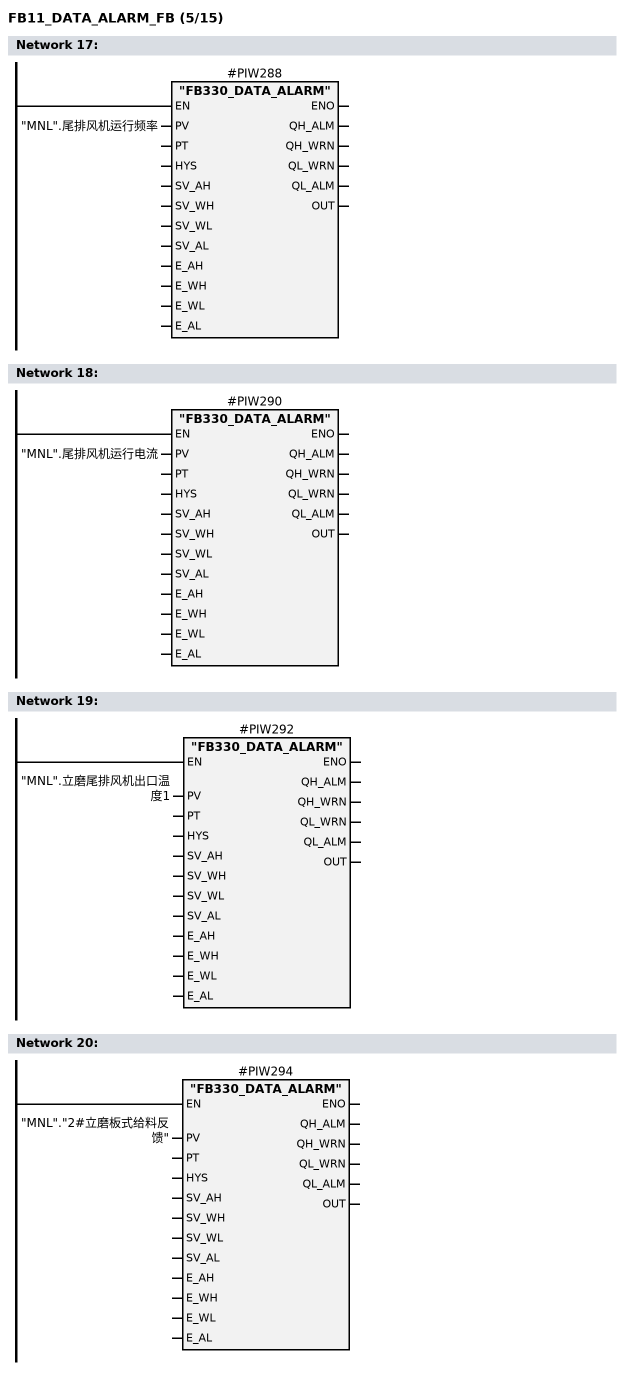
   RUNG wire#powerrail
      #PIW288(PV := "MNL".尾排风机运行频率, PT :=, HYS :=, SV_AH :=, SV_WH :=, SV_WL :=, SV_AL :=, E_AH :=, E_WH :=, E_WL :=, E_AL :=, QH_ALM =>, QH_WRN =>, QL_WRN =>, QL_ALM =>, OUT =>)
   END_RUNG
   // the same network as SCL:
   #PIW288(PV := "MNL".尾排风机运行频率);   // "FB330_DATA_ALARM"
END_REGION

REGION Network 18
   RUNG wire#powerrail
      #PIW290(PV := "MNL".尾排风机运行电流, PT :=, HYS :=, SV_AH :=, SV_WH :=, SV_WL :=, SV_AL :=, E_AH :=, E_WH :=, E_WL :=, E_AL :=, QH_ALM =>, QH_WRN =>, QL_WRN =>, QL_ALM =>, OUT =>)
   END_RUNG
   // the same network as SCL:
   #PIW290(PV := "MNL".尾排风机运行电流);   // "FB330_DATA_ALARM"
END_REGION

REGION Network 19
   RUNG wire#powerrail
      #PIW292(PV := "MNL".立磨尾排风机出口温度1, PT :=, HYS :=, SV_AH :=, SV_WH :=, SV_WL :=, SV_AL :=, E_AH :=, E_WH :=, E_WL :=, E_AL :=, QH_ALM =>, QH_WRN =>, QL_WRN =>, QL_ALM =>, OUT =>)
   END_RUNG
   // the same network as SCL:
   #PIW292(PV := "MNL".立磨尾排风机出口温度1);   // "FB330_DATA_ALARM"
END_REGION

REGION Network 20
   RUNG wire#powerrail
      #PIW294(PV := "MNL"."2#立磨板式给料反馈", PT :=, HYS :=, SV_AH :=, SV_WH :=, SV_WL :=, SV_AL :=, E_AH :=, E_WH :=, E_WL :=, E_AL :=, QH_ALM =>, QH_WRN =>, QL_WRN =>, QL_ALM =>, OUT =>)
   END_RUNG
   // the same network as SCL:
   #PIW294(PV := "MNL"."2#立磨板式给料反馈");   // "FB330_DATA_ALARM"
END_REGION

REGION Network 21
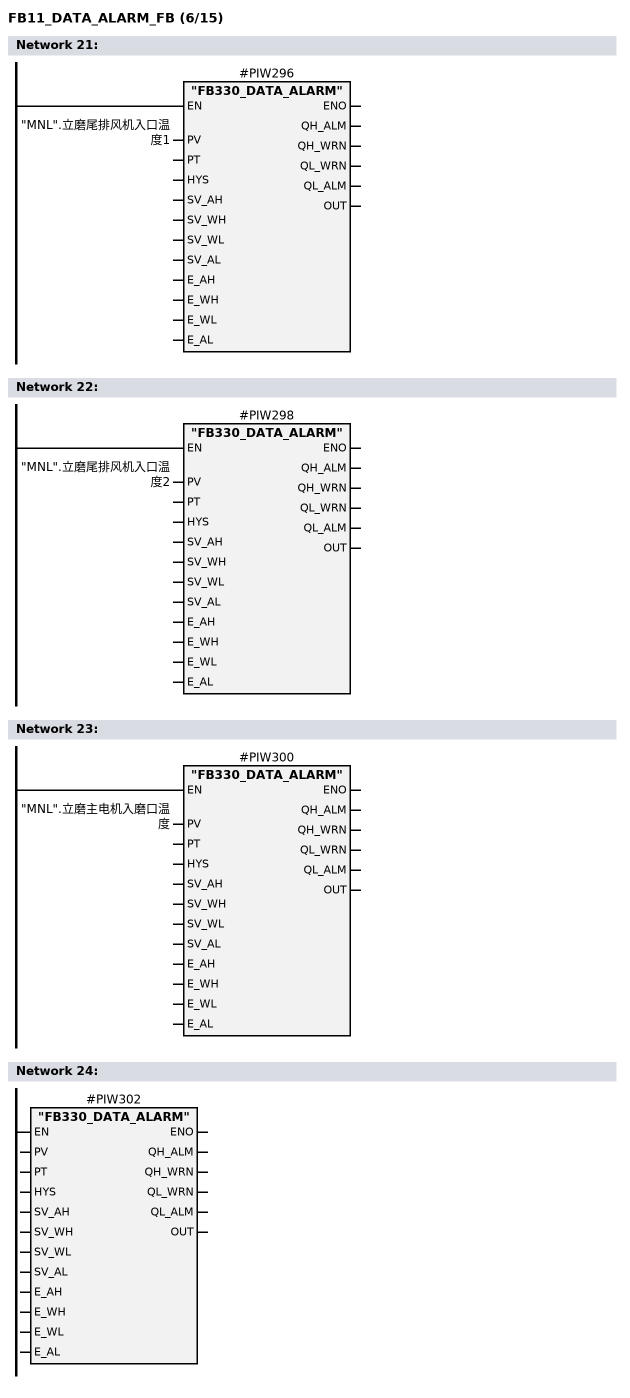
   RUNG wire#powerrail
      #PIW296(PV := "MNL".立磨尾排风机入口温度1, PT :=, HYS :=, SV_AH :=, SV_WH :=, SV_WL :=, SV_AL :=, E_AH :=, E_WH :=, E_WL :=, E_AL :=, QH_ALM =>, QH_WRN =>, QL_WRN =>, QL_ALM =>, OUT =>)
   END_RUNG
   // the same network as SCL:
   #PIW296(PV := "MNL".立磨尾排风机入口温度1);   // "FB330_DATA_ALARM"
END_REGION

REGION Network 22
   RUNG wire#powerrail
      #PIW298(PV := "MNL".立磨尾排风机入口温度2, PT :=, HYS :=, SV_AH :=, SV_WH :=, SV_WL :=, SV_AL :=, E_AH :=, E_WH :=, E_WL :=, E_AL :=, QH_ALM =>, QH_WRN =>, QL_WRN =>, QL_ALM =>, OUT =>)
   END_RUNG
   // the same network as SCL:
   #PIW298(PV := "MNL".立磨尾排风机入口温度2);   // "FB330_DATA_ALARM"
END_REGION

REGION Network 23
   RUNG wire#powerrail
      #PIW300(PV := "MNL".立磨主电机入磨口温度, PT :=, HYS :=, SV_AH :=, SV_WH :=, SV_WL :=, SV_AL :=, E_AH :=, E_WH :=, E_WL :=, E_AL :=, QH_ALM =>, QH_WRN =>, QL_WRN =>, QL_ALM =>, OUT =>)
   END_RUNG
   // the same network as SCL:
   #PIW300(PV := "MNL".立磨主电机入磨口温度);   // "FB330_DATA_ALARM"
END_REGION

REGION Network 24
   RUNG wire#powerrail
      #PIW302(PV :=, PT :=, HYS :=, SV_AH :=, SV_WH :=, SV_WL :=, SV_AL :=, E_AH :=, E_WH :=, E_WL :=, E_AL :=, QH_ALM =>, QH_WRN =>, QL_WRN =>, QL_ALM =>, OUT =>)
   END_RUNG
   // the same network as SCL:
   #PIW302();   // "FB330_DATA_ALARM"
END_REGION

REGION Network 25
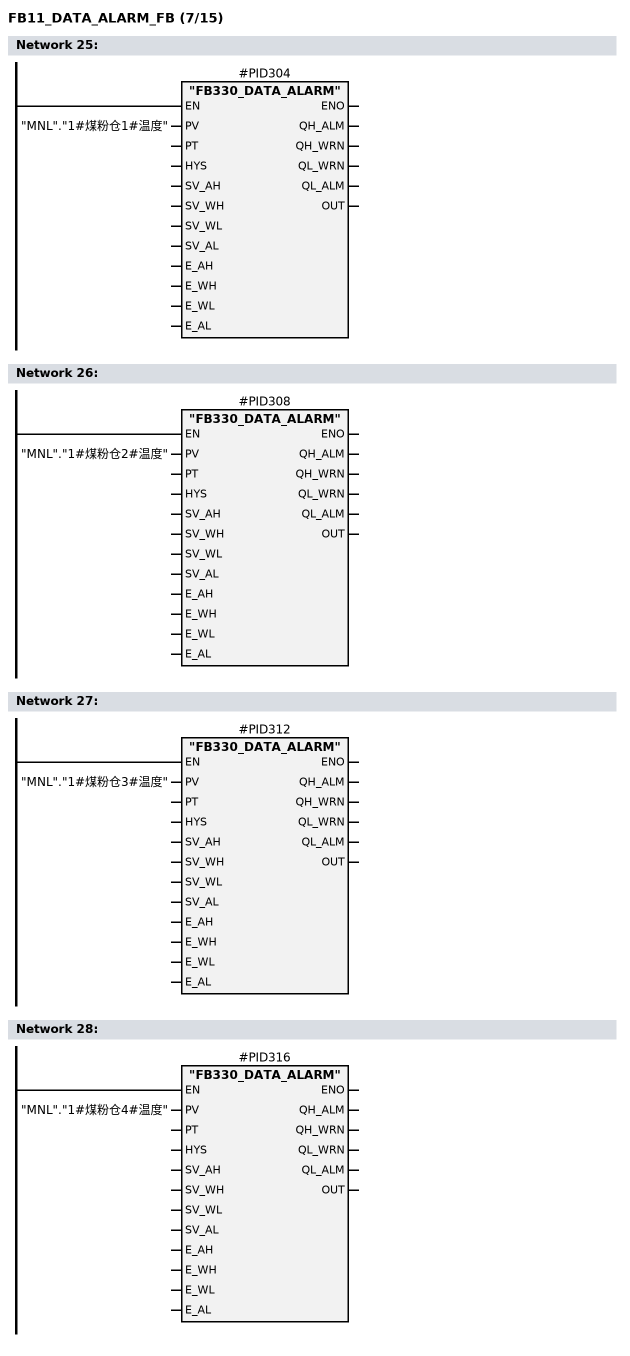
   RUNG wire#powerrail
      #PID304(PV := "MNL"."1#煤粉仓1#温度", PT :=, HYS :=, SV_AH :=, SV_WH :=, SV_WL :=, SV_AL :=, E_AH :=, E_WH :=, E_WL :=, E_AL :=, QH_ALM =>, QH_WRN =>, QL_WRN =>, QL_ALM =>, OUT =>)
   END_RUNG
   // the same network as SCL:
   #PID304(PV := "MNL"."1#煤粉仓1#温度");   // "FB330_DATA_ALARM"
END_REGION

REGION Network 26
   RUNG wire#powerrail
      #PID308(PV := "MNL"."1#煤粉仓2#温度", PT :=, HYS :=, SV_AH :=, SV_WH :=, SV_WL :=, SV_AL :=, E_AH :=, E_WH :=, E_WL :=, E_AL :=, QH_ALM =>, QH_WRN =>, QL_WRN =>, QL_ALM =>, OUT =>)
   END_RUNG
   // the same network as SCL:
   #PID308(PV := "MNL"."1#煤粉仓2#温度");   // "FB330_DATA_ALARM"
END_REGION

REGION Network 27
   RUNG wire#powerrail
      #PID312(PV := "MNL"."1#煤粉仓3#温度", PT :=, HYS :=, SV_AH :=, SV_WH :=, SV_WL :=, SV_AL :=, E_AH :=, E_WH :=, E_WL :=, E_AL :=, QH_ALM =>, QH_WRN =>, QL_WRN =>, QL_ALM =>, OUT =>)
   END_RUNG
   // the same network as SCL:
   #PID312(PV := "MNL"."1#煤粉仓3#温度");   // "FB330_DATA_ALARM"
END_REGION

REGION Network 28
   RUNG wire#powerrail
      #PID316(PV := "MNL"."1#煤粉仓4#温度", PT :=, HYS :=, SV_AH :=, SV_WH :=, SV_WL :=, SV_AL :=, E_AH :=, E_WH :=, E_WL :=, E_AL :=, QH_ALM =>, QH_WRN =>, QL_WRN =>, QL_ALM =>, OUT =>)
   END_RUNG
   // the same network as SCL:
   #PID316(PV := "MNL"."1#煤粉仓4#温度");   // "FB330_DATA_ALARM"
END_REGION

REGION Network 29
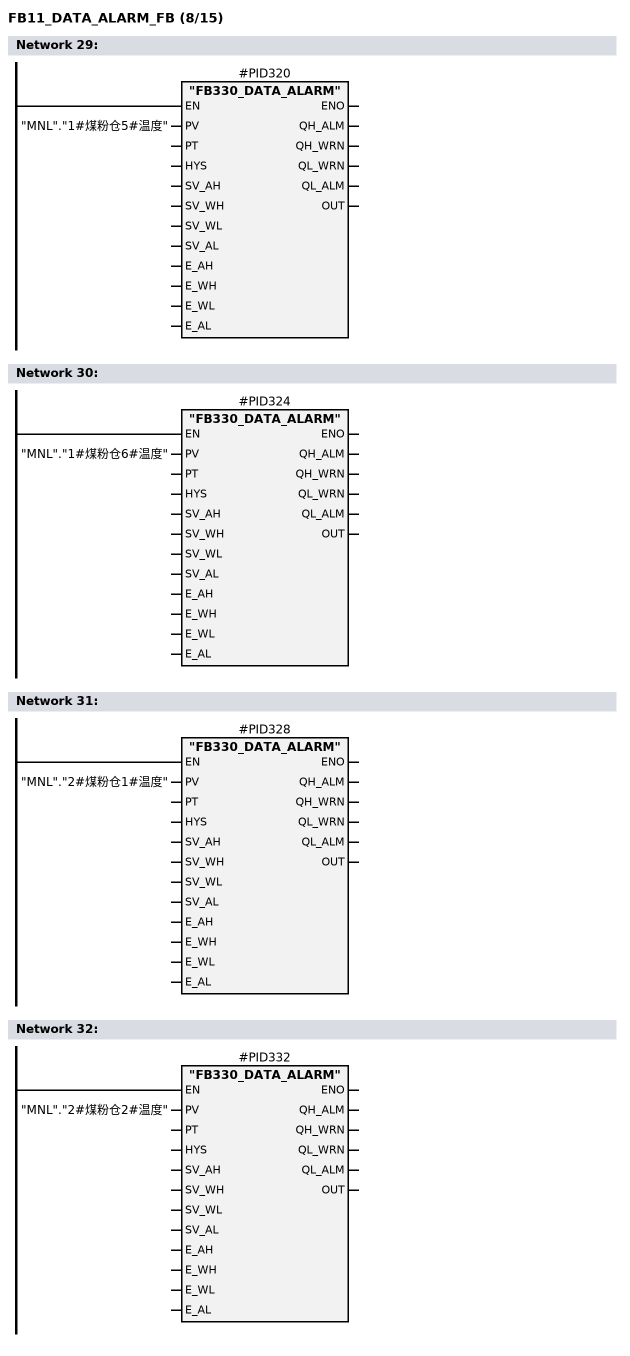
   RUNG wire#powerrail
      #PID320(PV := "MNL"."1#煤粉仓5#温度", PT :=, HYS :=, SV_AH :=, SV_WH :=, SV_WL :=, SV_AL :=, E_AH :=, E_WH :=, E_WL :=, E_AL :=, QH_ALM =>, QH_WRN =>, QL_WRN =>, QL_ALM =>, OUT =>)
   END_RUNG
   // the same network as SCL:
   #PID320(PV := "MNL"."1#煤粉仓5#温度");   // "FB330_DATA_ALARM"
END_REGION

REGION Network 30
   RUNG wire#powerrail
      #PID324(PV := "MNL"."1#煤粉仓6#温度", PT :=, HYS :=, SV_AH :=, SV_WH :=, SV_WL :=, SV_AL :=, E_AH :=, E_WH :=, E_WL :=, E_AL :=, QH_ALM =>, QH_WRN =>, QL_WRN =>, QL_ALM =>, OUT =>)
   END_RUNG
   // the same network as SCL:
   #PID324(PV := "MNL"."1#煤粉仓6#温度");   // "FB330_DATA_ALARM"
END_REGION

REGION Network 31
   RUNG wire#powerrail
      #PID328(PV := "MNL"."2#煤粉仓1#温度", PT :=, HYS :=, SV_AH :=, SV_WH :=, SV_WL :=, SV_AL :=, E_AH :=, E_WH :=, E_WL :=, E_AL :=, QH_ALM =>, QH_WRN =>, QL_WRN =>, QL_ALM =>, OUT =>)
   END_RUNG
   // the same network as SCL:
   #PID328(PV := "MNL"."2#煤粉仓1#温度");   // "FB330_DATA_ALARM"
END_REGION

REGION Network 32
   RUNG wire#powerrail
      #PID332(PV := "MNL"."2#煤粉仓2#温度", PT :=, HYS :=, SV_AH :=, SV_WH :=, SV_WL :=, SV_AL :=, E_AH :=, E_WH :=, E_WL :=, E_AL :=, QH_ALM =>, QH_WRN =>, QL_WRN =>, QL_ALM =>, OUT =>)
   END_RUNG
   // the same network as SCL:
   #PID332(PV := "MNL"."2#煤粉仓2#温度");   // "FB330_DATA_ALARM"
END_REGION

REGION Network 33
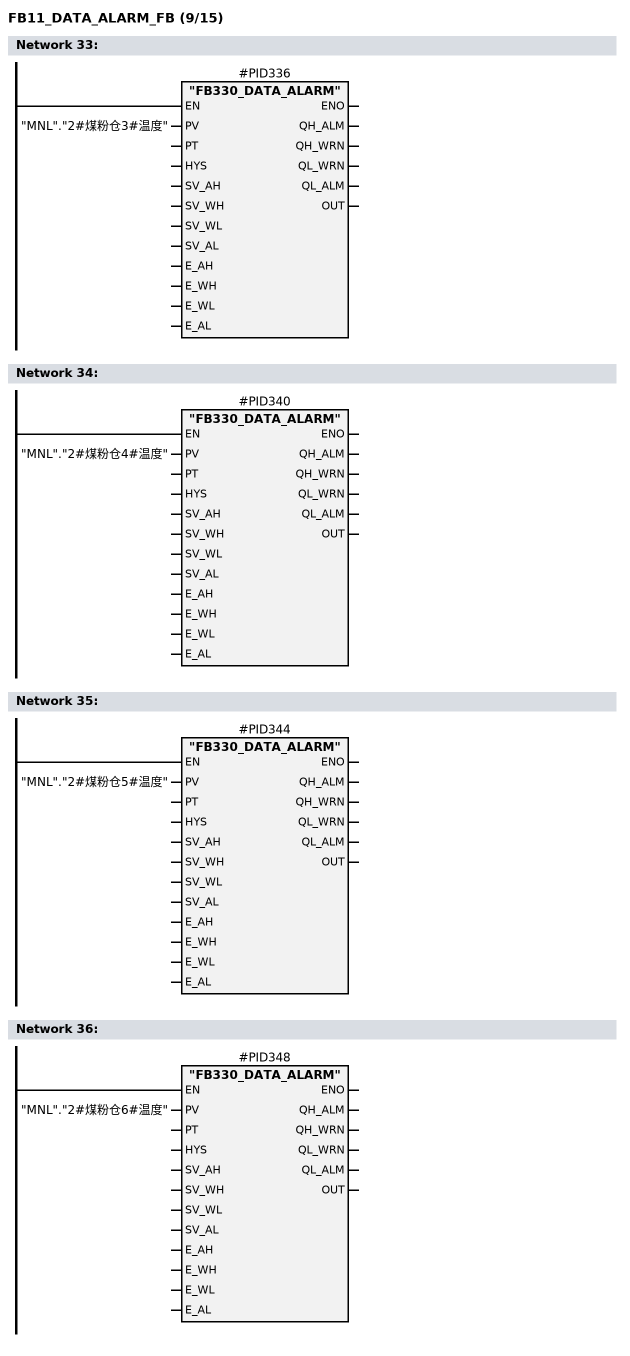
   RUNG wire#powerrail
      #PID336(PV := "MNL"."2#煤粉仓3#温度", PT :=, HYS :=, SV_AH :=, SV_WH :=, SV_WL :=, SV_AL :=, E_AH :=, E_WH :=, E_WL :=, E_AL :=, QH_ALM =>, QH_WRN =>, QL_WRN =>, QL_ALM =>, OUT =>)
   END_RUNG
   // the same network as SCL:
   #PID336(PV := "MNL"."2#煤粉仓3#温度");   // "FB330_DATA_ALARM"
END_REGION

REGION Network 34
   RUNG wire#powerrail
      #PID340(PV := "MNL"."2#煤粉仓4#温度", PT :=, HYS :=, SV_AH :=, SV_WH :=, SV_WL :=, SV_AL :=, E_AH :=, E_WH :=, E_WL :=, E_AL :=, QH_ALM =>, QH_WRN =>, QL_WRN =>, QL_ALM =>, OUT =>)
   END_RUNG
   // the same network as SCL:
   #PID340(PV := "MNL"."2#煤粉仓4#温度");   // "FB330_DATA_ALARM"
END_REGION

REGION Network 35
   RUNG wire#powerrail
      #PID344(PV := "MNL"."2#煤粉仓5#温度", PT :=, HYS :=, SV_AH :=, SV_WH :=, SV_WL :=, SV_AL :=, E_AH :=, E_WH :=, E_WL :=, E_AL :=, QH_ALM =>, QH_WRN =>, QL_WRN =>, QL_ALM =>, OUT =>)
   END_RUNG
   // the same network as SCL:
   #PID344(PV := "MNL"."2#煤粉仓5#温度");   // "FB330_DATA_ALARM"
END_REGION

REGION Network 36
   RUNG wire#powerrail
      #PID348(PV := "MNL"."2#煤粉仓6#温度", PT :=, HYS :=, SV_AH :=, SV_WH :=, SV_WL :=, SV_AL :=, E_AH :=, E_WH :=, E_WL :=, E_AL :=, QH_ALM =>, QH_WRN =>, QL_WRN =>, QL_ALM =>, OUT =>)
   END_RUNG
   // the same network as SCL:
   #PID348(PV := "MNL"."2#煤粉仓6#温度");   // "FB330_DATA_ALARM"
END_REGION

REGION Network 37
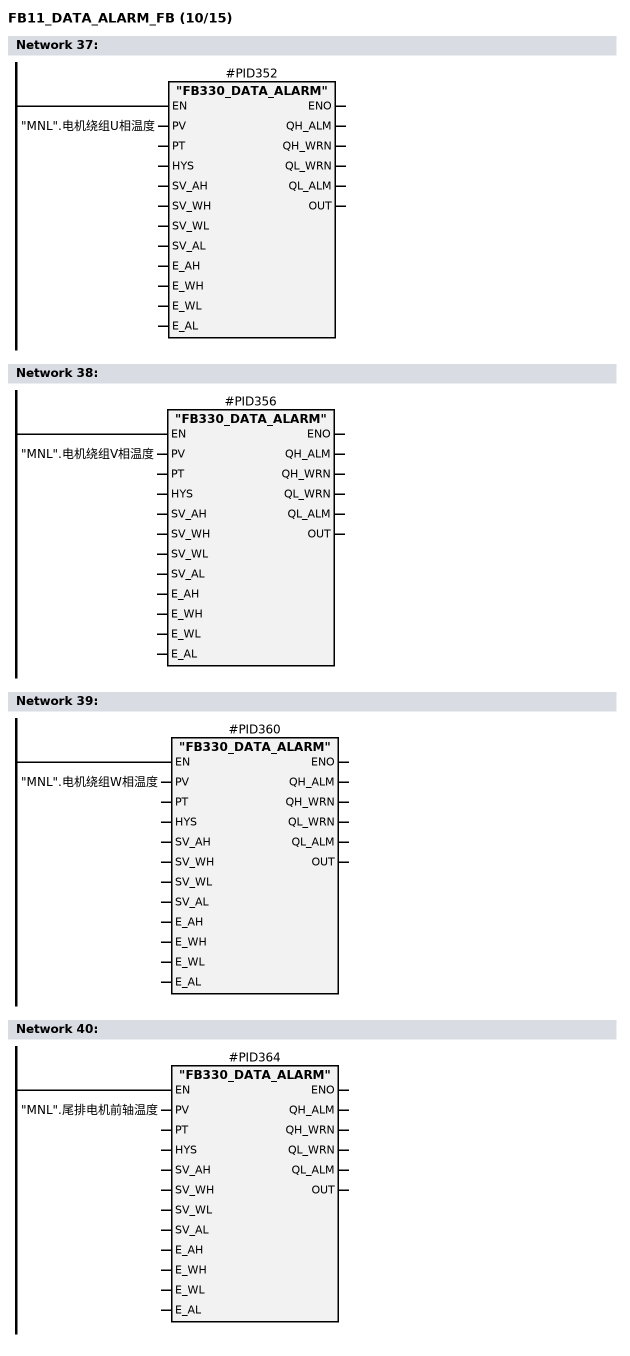
   RUNG wire#powerrail
      #PID352(PV := "MNL".电机绕组U相温度, PT :=, HYS :=, SV_AH :=, SV_WH :=, SV_WL :=, SV_AL :=, E_AH :=, E_WH :=, E_WL :=, E_AL :=, QH_ALM =>, QH_WRN =>, QL_WRN =>, QL_ALM =>, OUT =>)
   END_RUNG
   // the same network as SCL:
   #PID352(PV := "MNL".电机绕组U相温度);   // "FB330_DATA_ALARM"
END_REGION

REGION Network 38
   RUNG wire#powerrail
      #PID356(PV := "MNL".电机绕组V相温度, PT :=, HYS :=, SV_AH :=, SV_WH :=, SV_WL :=, SV_AL :=, E_AH :=, E_WH :=, E_WL :=, E_AL :=, QH_ALM =>, QH_WRN =>, QL_WRN =>, QL_ALM =>, OUT =>)
   END_RUNG
   // the same network as SCL:
   #PID356(PV := "MNL".电机绕组V相温度);   // "FB330_DATA_ALARM"
END_REGION

REGION Network 39
   RUNG wire#powerrail
      #PID360(PV := "MNL".电机绕组W相温度, PT :=, HYS :=, SV_AH :=, SV_WH :=, SV_WL :=, SV_AL :=, E_AH :=, E_WH :=, E_WL :=, E_AL :=, QH_ALM =>, QH_WRN =>, QL_WRN =>, QL_ALM =>, OUT =>)
   END_RUNG
   // the same network as SCL:
   #PID360(PV := "MNL".电机绕组W相温度);   // "FB330_DATA_ALARM"
END_REGION

REGION Network 40
   RUNG wire#powerrail
      #PID364(PV := "MNL".尾排电机前轴温度, PT :=, HYS :=, SV_AH :=, SV_WH :=, SV_WL :=, SV_AL :=, E_AH :=, E_WH :=, E_WL :=, E_AL :=, QH_ALM =>, QH_WRN =>, QL_WRN =>, QL_ALM =>, OUT =>)
   END_RUNG
   // the same network as SCL:
   #PID364(PV := "MNL".尾排电机前轴温度);   // "FB330_DATA_ALARM"
END_REGION

REGION Network 41
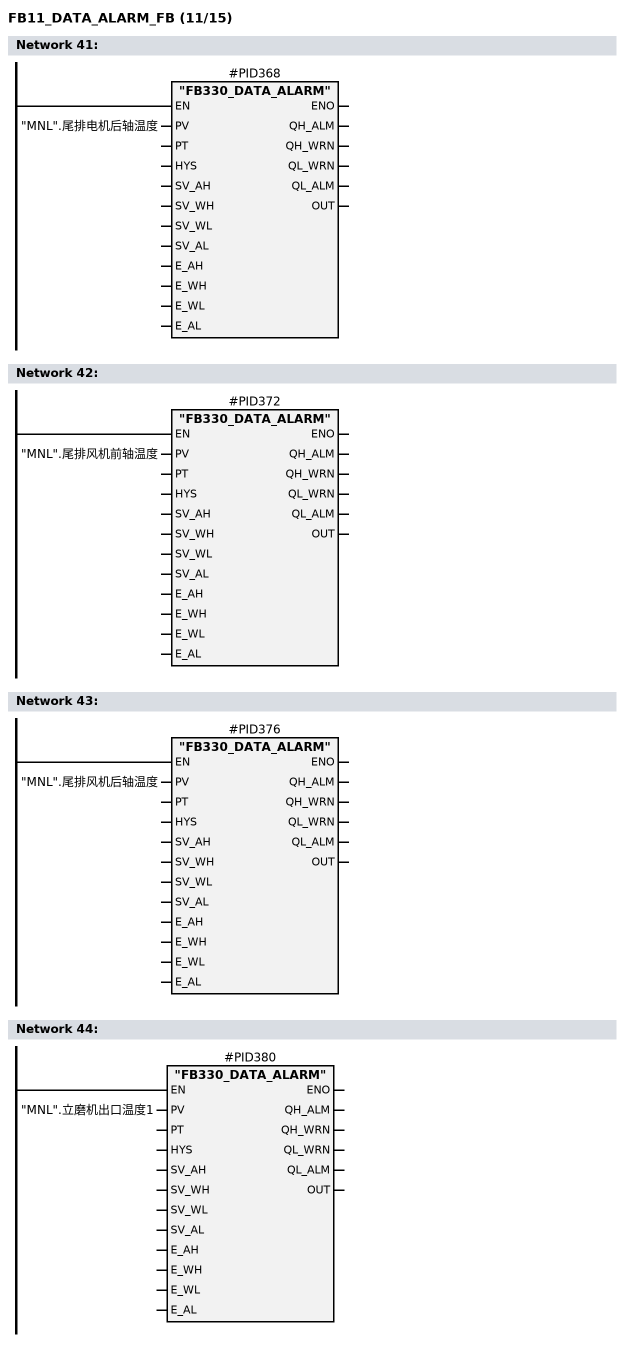
   RUNG wire#powerrail
      #PID368(PV := "MNL".尾排电机后轴温度, PT :=, HYS :=, SV_AH :=, SV_WH :=, SV_WL :=, SV_AL :=, E_AH :=, E_WH :=, E_WL :=, E_AL :=, QH_ALM =>, QH_WRN =>, QL_WRN =>, QL_ALM =>, OUT =>)
   END_RUNG
   // the same network as SCL:
   #PID368(PV := "MNL".尾排电机后轴温度);   // "FB330_DATA_ALARM"
END_REGION

REGION Network 42
   RUNG wire#powerrail
      #PID372(PV := "MNL".尾排风机前轴温度, PT :=, HYS :=, SV_AH :=, SV_WH :=, SV_WL :=, SV_AL :=, E_AH :=, E_WH :=, E_WL :=, E_AL :=, QH_ALM =>, QH_WRN =>, QL_WRN =>, QL_ALM =>, OUT =>)
   END_RUNG
   // the same network as SCL:
   #PID372(PV := "MNL".尾排风机前轴温度);   // "FB330_DATA_ALARM"
END_REGION

REGION Network 43
   RUNG wire#powerrail
      #PID376(PV := "MNL".尾排风机后轴温度, PT :=, HYS :=, SV_AH :=, SV_WH :=, SV_WL :=, SV_AL :=, E_AH :=, E_WH :=, E_WL :=, E_AL :=, QH_ALM =>, QH_WRN =>, QL_WRN =>, QL_ALM =>, OUT =>)
   END_RUNG
   // the same network as SCL:
   #PID376(PV := "MNL".尾排风机后轴温度);   // "FB330_DATA_ALARM"
END_REGION

REGION Network 44
   RUNG wire#powerrail
      #PID380(PV := "MNL".立磨机出口温度1, PT :=, HYS :=, SV_AH :=, SV_WH :=, SV_WL :=, SV_AL :=, E_AH :=, E_WH :=, E_WL :=, E_AL :=, QH_ALM =>, QH_WRN =>, QL_WRN =>, QL_ALM =>, OUT =>)
   END_RUNG
   // the same network as SCL:
   #PID380(PV := "MNL".立磨机出口温度1);   // "FB330_DATA_ALARM"
END_REGION

REGION Network 45
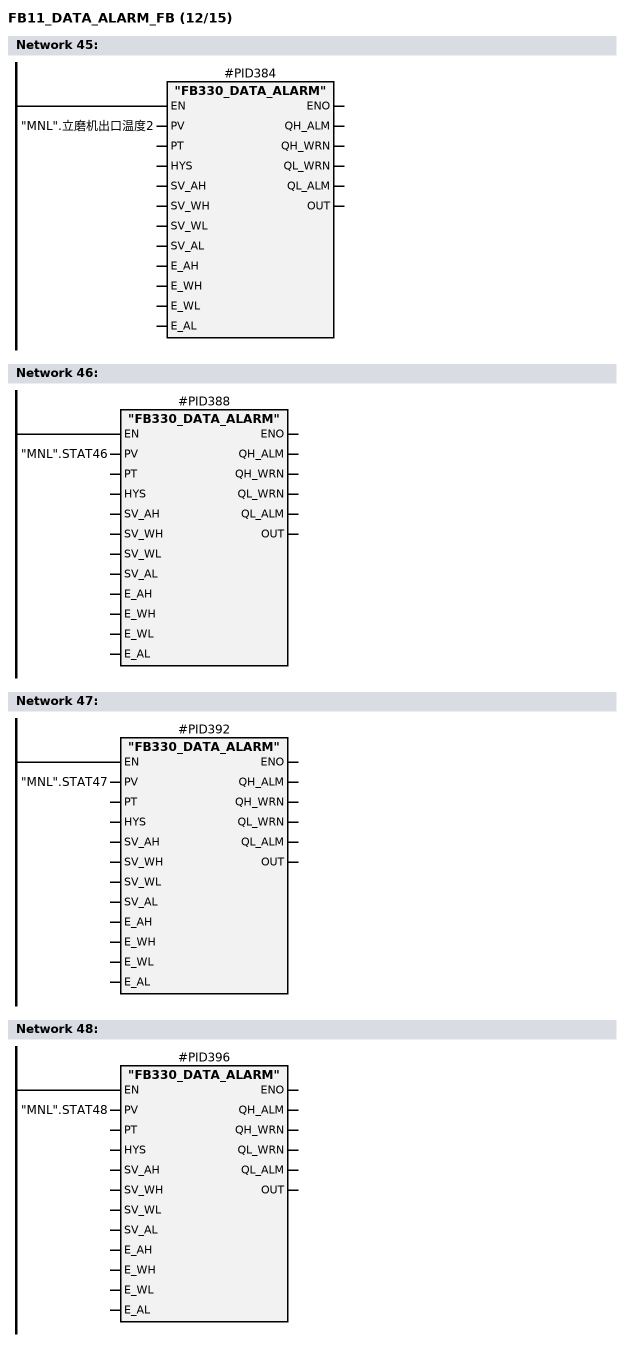
   RUNG wire#powerrail
      #PID384(PV := "MNL".立磨机出口温度2, PT :=, HYS :=, SV_AH :=, SV_WH :=, SV_WL :=, SV_AL :=, E_AH :=, E_WH :=, E_WL :=, E_AL :=, QH_ALM =>, QH_WRN =>, QL_WRN =>, QL_ALM =>, OUT =>)
   END_RUNG
   // the same network as SCL:
   #PID384(PV := "MNL".立磨机出口温度2);   // "FB330_DATA_ALARM"
END_REGION

REGION Network 46
   RUNG wire#powerrail
      #PID388(PV := "MNL".STAT46, PT :=, HYS :=, SV_AH :=, SV_WH :=, SV_WL :=, SV_AL :=, E_AH :=, E_WH :=, E_WL :=, E_AL :=, QH_ALM =>, QH_WRN =>, QL_WRN =>, QL_ALM =>, OUT =>)
   END_RUNG
   // the same network as SCL:
   #PID388(PV := "MNL".STAT46);   // "FB330_DATA_ALARM"
END_REGION

REGION Network 47
   RUNG wire#powerrail
      #PID392(PV := "MNL".STAT47, PT :=, HYS :=, SV_AH :=, SV_WH :=, SV_WL :=, SV_AL :=, E_AH :=, E_WH :=, E_WL :=, E_AL :=, QH_ALM =>, QH_WRN =>, QL_WRN =>, QL_ALM =>, OUT =>)
   END_RUNG
   // the same network as SCL:
   #PID392(PV := "MNL".STAT47);   // "FB330_DATA_ALARM"
END_REGION

REGION Network 48
   RUNG wire#powerrail
      #PID396(PV := "MNL".STAT48, PT :=, HYS :=, SV_AH :=, SV_WH :=, SV_WL :=, SV_AL :=, E_AH :=, E_WH :=, E_WL :=, E_AL :=, QH_ALM =>, QH_WRN =>, QL_WRN =>, QL_ALM =>, OUT =>)
   END_RUNG
   // the same network as SCL:
   #PID396(PV := "MNL".STAT48);   // "FB330_DATA_ALARM"
END_REGION

REGION Network 49
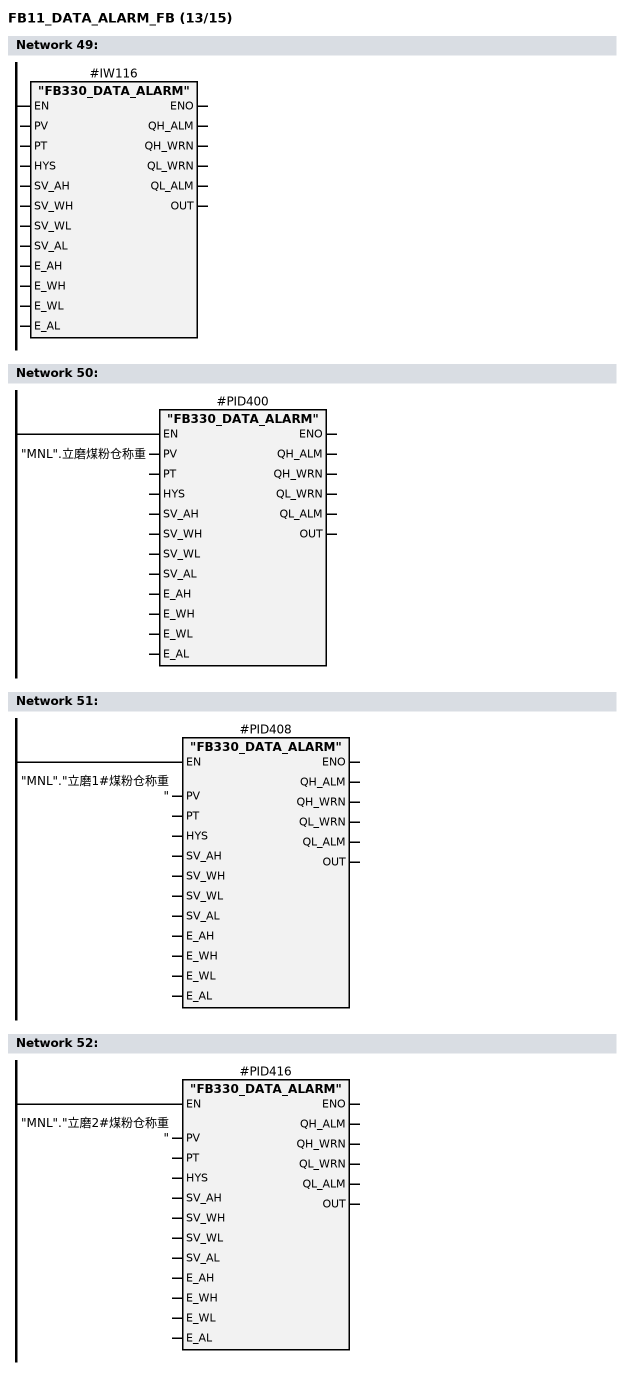
   RUNG wire#powerrail
      #IW116(PV :=, PT :=, HYS :=, SV_AH :=, SV_WH :=, SV_WL :=, SV_AL :=, E_AH :=, E_WH :=, E_WL :=, E_AL :=, QH_ALM =>, QH_WRN =>, QL_WRN =>, QL_ALM =>, OUT =>)
   END_RUNG
   // the same network as SCL:
   #IW116();   // "FB330_DATA_ALARM"
END_REGION

REGION Network 50
   RUNG wire#powerrail
      #PID400(PV := "MNL".立磨煤粉仓称重, PT :=, HYS :=, SV_AH :=, SV_WH :=, SV_WL :=, SV_AL :=, E_AH :=, E_WH :=, E_WL :=, E_AL :=, QH_ALM =>, QH_WRN =>, QL_WRN =>, QL_ALM =>, OUT =>)
   END_RUNG
   // the same network as SCL:
   #PID400(PV := "MNL".立磨煤粉仓称重);   // "FB330_DATA_ALARM"
END_REGION

REGION Network 51
   RUNG wire#powerrail
      #PID408(PV := "MNL"."立磨1#煤粉仓称重", PT :=, HYS :=, SV_AH :=, SV_WH :=, SV_WL :=, SV_AL :=, E_AH :=, E_WH :=, E_WL :=, E_AL :=, QH_ALM =>, QH_WRN =>, QL_WRN =>, QL_ALM =>, OUT =>)
   END_RUNG
   // the same network as SCL:
   #PID408(PV := "MNL"."立磨1#煤粉仓称重");   // "FB330_DATA_ALARM"
END_REGION

REGION Network 52
   RUNG wire#powerrail
      #PID416(PV := "MNL"."立磨2#煤粉仓称重", PT :=, HYS :=, SV_AH :=, SV_WH :=, SV_WL :=, SV_AL :=, E_AH :=, E_WH :=, E_WL :=, E_AL :=, QH_ALM =>, QH_WRN =>, QL_WRN =>, QL_ALM =>, OUT =>)
   END_RUNG
   // the same network as SCL:
   #PID416(PV := "MNL"."立磨2#煤粉仓称重");   // "FB330_DATA_ALARM"
END_REGION

REGION Network 53
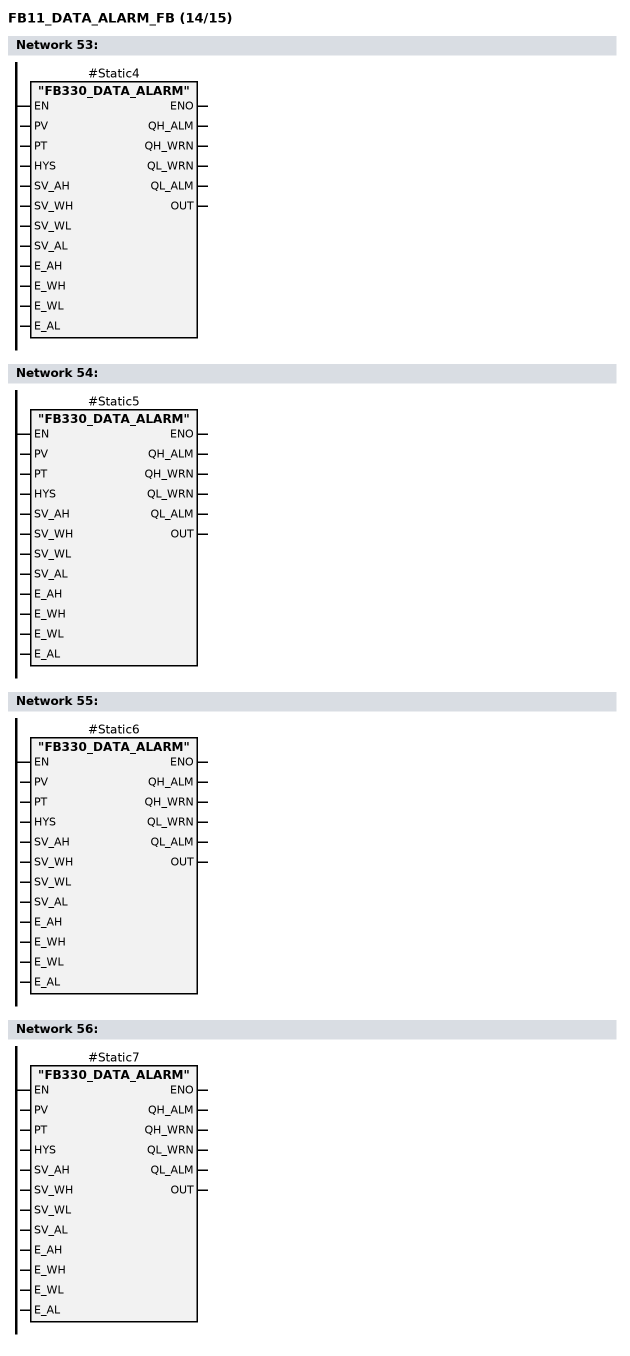
   RUNG wire#powerrail
      #Static4(PV :=, PT :=, HYS :=, SV_AH :=, SV_WH :=, SV_WL :=, SV_AL :=, E_AH :=, E_WH :=, E_WL :=, E_AL :=, QH_ALM =>, QH_WRN =>, QL_WRN =>, QL_ALM =>, OUT =>)
   END_RUNG
   // the same network as SCL:
   #Static4();   // "FB330_DATA_ALARM"
END_REGION

REGION Network 54
   RUNG wire#powerrail
      #Static5(PV :=, PT :=, HYS :=, SV_AH :=, SV_WH :=, SV_WL :=, SV_AL :=, E_AH :=, E_WH :=, E_WL :=, E_AL :=, QH_ALM =>, QH_WRN =>, QL_WRN =>, QL_ALM =>, OUT =>)
   END_RUNG
   // the same network as SCL:
   #Static5();   // "FB330_DATA_ALARM"
END_REGION

REGION Network 55
   RUNG wire#powerrail
      #Static6(PV :=, PT :=, HYS :=, SV_AH :=, SV_WH :=, SV_WL :=, SV_AL :=, E_AH :=, E_WH :=, E_WL :=, E_AL :=, QH_ALM =>, QH_WRN =>, QL_WRN =>, QL_ALM =>, OUT =>)
   END_RUNG
   // the same network as SCL:
   #Static6();   // "FB330_DATA_ALARM"
END_REGION

REGION Network 56
   RUNG wire#powerrail
      #Static7(PV :=, PT :=, HYS :=, SV_AH :=, SV_WH :=, SV_WL :=, SV_AL :=, E_AH :=, E_WH :=, E_WL :=, E_AL :=, QH_ALM =>, QH_WRN =>, QL_WRN =>, QL_ALM =>, OUT =>)
   END_RUNG
   // the same network as SCL:
   #Static7();   // "FB330_DATA_ALARM"
END_REGION

REGION Network 57
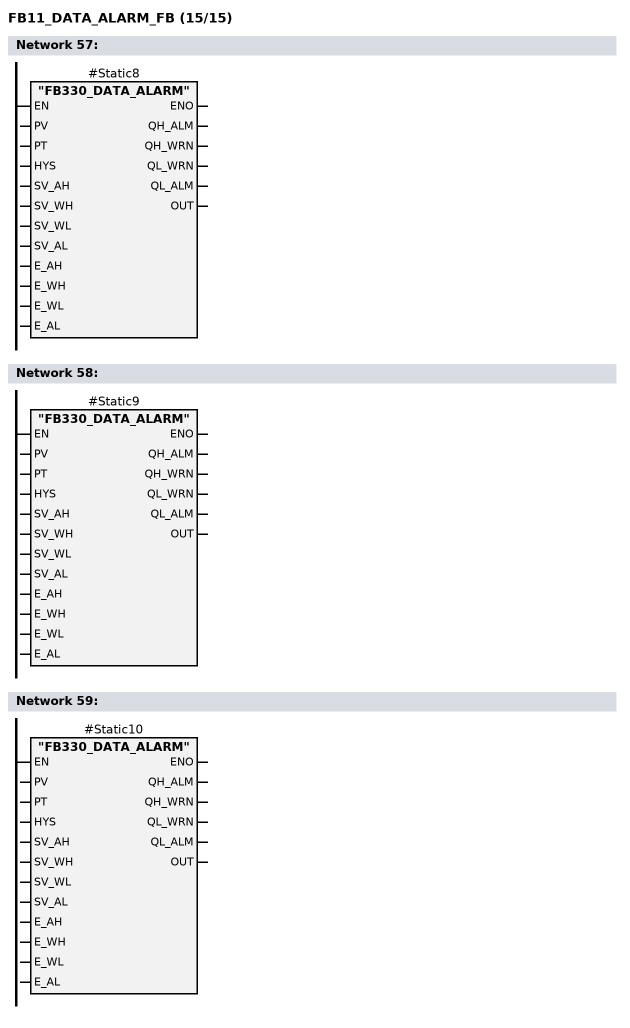
   RUNG wire#powerrail
      #Static8(PV :=, PT :=, HYS :=, SV_AH :=, SV_WH :=, SV_WL :=, SV_AL :=, E_AH :=, E_WH :=, E_WL :=, E_AL :=, QH_ALM =>, QH_WRN =>, QL_WRN =>, QL_ALM =>, OUT =>)
   END_RUNG
   // the same network as SCL:
   #Static8();   // "FB330_DATA_ALARM"
END_REGION

REGION Network 58
   RUNG wire#powerrail
      #Static9(PV :=, PT :=, HYS :=, SV_AH :=, SV_WH :=, SV_WL :=, SV_AL :=, E_AH :=, E_WH :=, E_WL :=, E_AL :=, QH_ALM =>, QH_WRN =>, QL_WRN =>, QL_ALM =>, OUT =>)
   END_RUNG
   // the same network as SCL:
   #Static9();   // "FB330_DATA_ALARM"
END_REGION

REGION Network 59
   RUNG wire#powerrail
      #Static10(PV :=, PT :=, HYS :=, SV_AH :=, SV_WH :=, SV_WL :=, SV_AL :=, E_AH :=, E_WH :=, E_WL :=, E_AL :=, QH_ALM =>, QH_WRN =>, QL_WRN =>, QL_ALM =>, OUT =>)
   END_RUNG
   // the same network as SCL:
   #Static10();   // "FB330_DATA_ALARM"
END_REGION
END_FUNCTION_BLOCK

FUNCTION_BLOCK "阀门控制块"   // FB300, LAD
{ S7_Optimized_Access := 'TRUE' }
VERSION : 0.1
   VAR_INPUT
      LR : Bool;
      V_OPEN : Bool;
      V_CLOSE : Bool;
      HMI_OPEN : Bool;
      HMI_CLOSE : Bool;
   END_VAR
   VAR_OUTPUT
      OUT_OP_PULSE : Bool;
      OUT_CL_PULSE : Bool;
   END_VAR
   VAR_IN_OUT
      OUT_HOLD : Bool;
   END_VAR
BEGIN

REGION Network 1
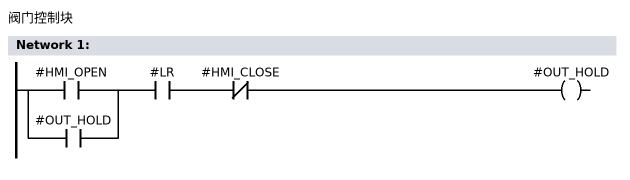
   RUNG wire#powerrail
      Contact( #HMI_OPEN )
      wire#w1
      Contact( #LR )
      I_Contact( #HMI_CLOSE )
      Coil( #OUT_HOLD )
   END_RUNG
   RUNG wire#powerrail
      Contact( #OUT_HOLD )
   END_RUNG wire#w1
   // the same network as SCL:
   #OUT_HOLD := (#HMI_OPEN OR #OUT_HOLD) AND #LR AND NOT #HMI_CLOSE;
END_REGION
END_FUNCTION_BLOCK

FUNCTION_BLOCK "FB330_DATA_ALARM"   // FB330, LAD
{ S7_Optimized_Access := 'FALSE' }
VERSION : 0.1
// REAL的报警块
   VAR_INPUT
      PV : Real;   // 过程值
      PT : Real := 1.0;   // 系数
      HYS : Real;   // 回差值
      SV_AH : Real;   // 高报警设定值
      SV_WH : Real;   // 高警告设定值
      SV_WL : Real;   // 低警告设定值
      SV_AL : Real;   // 低报警设定值
      E_AH : Bool;   // 高报警使能
      E_WH : Bool;   // 高警告使能
      E_WL : Bool;   // 低警告使能
      E_AL : Bool;   // 低报警使能
   END_VAR
   VAR_OUTPUT
      QH_ALM : Bool;   // 高报警输出
      QH_WRN : Bool;   // 高警告输出
      QL_WRN : Bool;   // 低警告输出
      QL_ALM : Bool;   // 低报警输出
      OUT : Real;   // 输出
   END_VAR
   VAR
      SR1 : Bool;
      SR2 : Bool;
      SR3 : Bool;
      SR4 : Bool;
   END_VAR
   VAR_TEMP
      TEMP_AH : Real;
      TEMP_WH : Real;
      TEMP_AL : Real;
      TEMP_WL : Real;
      TEMP_OUT : Real;
   END_VAR
BEGIN

REGION Network 1
   // 系数转换
